   "PLC_a_HMI_Fila[6].Elemento[2].Estado" : Byte, 100 ms
   "PLC_a_HMI_Fila[6].Elemento[3].Figura" : Byte, 100 ms
   "PLC_a_HMI_Fila[6].Elemento[3].Offset_X" : Int, 100 ms
   "PLC_a_HMI_Fila[6].Elemento[3].Estado" : Byte, 100 ms
   "PLC_a_HMI_Fila[6].Elemento[4].Figura" : Byte, 100 ms
   "PLC_a_HMI_Fila[6].Elemento[4].Offset_X" : Int, 100 ms
   "PLC_a_HMI_Fila[6].Elemento[4].Estado" : Byte, 100 ms
   "PLC_a_HMI_Fila[6].Elemento[5].Figura" : Byte, 100 ms
   "PLC_a_HMI_Fila[6].Elemento[5].Offset_X" : Int, 100 ms
   "PLC_a_HMI_Fila[6].Elemento[5].Estado" : Byte, 100 ms
   "PLC_a_HMI_Fila[6].Elemento[6].Figura" : Byte, 100 ms
   "PLC_a_HMI_Fila[6].Elemento[6].Offset_X" : Int, 100 ms
   "PLC_a_HMI_Fila[6].Elemento[6].Estado" : Byte, 100 ms
   "PLC_a_HMI_Fila[6].Elemento[7].Figura" : Byte, 100 ms
   "PLC_a_HMI_Fila[6].Elemento[7].Offset_X" : Int, 100 ms
   "PLC_a_HMI_Fila[6].Elemento[7].Estado" : Byte, 100 ms
   "PLC_a_HMI_Fila[6].Elemento[8].Figura" : Byte, 100 ms
   "PLC_a_HMI_Fila[6].Elemento[8].Offset_X" : Int, 100 ms
   "PLC_a_HMI_Fila[6].Elemento[8].Estado" : Byte, 100 ms
   "PLC_a_HMI_Fila[6].Elemento[9].Figura" : Byte, 100 ms
   "PLC_a_HMI_Fila[6].Elemento[9].Offset_X" : Int, 100 ms
   "PLC_a_HMI_Fila[6].Elemento[9].Estado" : Byte, 100 ms
   "PLC_a_HMI_Fila[6].Elemento[10].Figura" : Byte, 100 ms
   "PLC_a_HMI_Fila[6].Elemento[10].Offset_X" : Int, 100 ms
   "PLC_a_HMI_Fila[6].Elemento[10].Estado" : Byte, 100 ms
   "PLC_a_HMI_Fila_Activa" : Byte, 1 s
   "DB_Animación_Figura_SEL" : Byte, 1 s
   "PLC_FechaHora" : Date_And_Time, 1 s
   "Proceso Empujador_Capa_Actual" : Byte, 1 s
   "DB_Receta_Actual_Nro_Capas_Pallet" : Byte, 1 s
   "Proceso Dosificador_Cant_Cajas" : Word, 1 s
   "DB_Receta_Actual_Nombre" : Array [0..49] of Char, 1 s
   "Proceso CargaPallet_Cant_Pallets" : DInt, 1 s
   "Proceso Empujador_Cant_Cajas" : DInt, 1 s
   "PLC a HMI_TRANSPORTES_Hab" : Bool, 1 s
   "PLC a HMI_Seg_Entrada_Envol" : Bool, 1 s
   "PLC a HMI_Seg_Salida_Envol" : Bool, 1 s
   "PLC a HMI_oTranspPall1" : Bool, 1 s
   "PLC a HMI_oTranspPall2" : Bool, 1 s
   "PLC a HMI_oTranspPall3" : Bool, 1 s
   "PLC a HMI_oTranspPall3Freno" : Bool, 1 s
   "PLC a HMI_oTranspPall4" : Bool, 1 s
   "PLC a HMI_oTranspPall5" : Bool, 1 s
   "PLC a HMI_iBrazoPos_Envolv" : Bool, 1 s
   "PLC a HMI_oHabilMovBrazo_Envol" : Bool, 1 s
   "PLC a HMI_iCartZonaSeg" : Bool, 1 s
   "PLC a HMI_iCartAplicado" : Bool, 1 s
   "PLC a HMI_iCartConAlarm" : Bool, 1 s
   "PLC a HMI_oTomarCartón" : Bool, 1 s
   "PLC a HMI_oAplicarCartón" : Bool, 1 s
   "PLC a HMI_oPaleZonaSeg" : Bool, 1 s
   "PLC a HMI_oPaleSinAlarm" : Bool, 1 s
   "FuncNormalAlterado" : Bool, 1 s
   "Confirmacion1" : Bool, internal
   "Confirmacion2" : Bool, internal

HMI tags "HMI_a_PLC"
   "HMI_Pls_Inc_Elem" : Bool, 1 s
   "HMI_Pls_Dec_Elem" : Bool, 1 s
   "HMI_Pls_Elem_Der" : Bool, 1 s
   "HMI_Pls_Elem_Izq" : Bool, 1 s
   "HMI_Pls_Inc_Fila" : Bool, 1 s
   "HMI_Pls_Dec_Fila" : Bool, 1 s
   "HMI_Pls_Fila_Sup" : Bool, 1 s
   "HMI_Pls_Fila_Inf" : Bool, 1 s
   "HMI_Pls_New_Fila" : Bool, 1 s
   "HMI_Pls_New_Elem" : Bool, 1 s
   "HMI_Pls_Kill_Elem" : Bool, 1 s
   "HMI_Pls_WR_Receta" : Bool, 1 s
   "HMI_Pls_RD_Receta" : Bool, 1 s
   "HMI_Imagen_Actual" : Word, 100 ms
   "HMI_Pls_Inc_Receta" : Bool, 1 s
   "HMI_Pls_Dec_Receta" : Bool, 1 s
   "HMI_Pls_Inc_Capa" : Bool, 1 s
   "HMI_Pls_Dec_Capa" : Bool, 1 s
   "HMI_Pls_Elem_+" : Bool, 1 s
   "HMI_Pls_Elem_-" : Bool, 1 s
   "HMI_Pls_CargarReceta" : Bool, 1 s
   "HMI_Pls_TerminarPallet" : Bool, 1 s
   "HMI_Pls_ResetPallets" : Bool, 1 s
   "HMI_Pls_ResetCajas" : Bool, 1 s
   "HMI_Pls_SalirImagenIni" : Bool, 1 s
   "HMI_Pls_MarMan_Ramp1" : Bool, 1 s
   "HMI_Pls_MarMan_Rol1" : Bool, 1 s
   "HMI_Pls_MarMan_Ramp2" : Bool, 1 s
   "HMI_Pls_MarMan_Rol2" : Bool, 1 s
   "HMI_Hab_Cartonero" : Bool, 1 s

discrete alarms
   1: '', class Grave, trigger "ALARMAS_1" bit 0
   2: '', class Grave, trigger "ALARMAS_1" bit 1
   3: '', class Grave, trigger "ALARMAS_1" bit 2
   4: '', class Grave, trigger "ALARMAS_1" bit 3
   5: '', class Grave, trigger "ALARMAS_1" bit 4
   6: '', class Grave, trigger "ALARMAS_1" bit 5
   7: '', class Grave, trigger "ALARMAS_1" bit 6
   8: '', class Grave, trigger "ALARMAS_1" bit 7
   9: '', class General, trigger "ALARMAS_1" bit 8
   10: '', class General, trigger "ALARMAS_1" bit 9
   11: '', class General, trigger "ALARMAS_1" bit 10
   12: '', class General, trigger "ALARMAS_1" bit 11
   13: '', class General, trigger "ALARMAS_1" bit 12
   14: '', class General, trigger "ALARMAS_1" bit 13
   15: '', class General, trigger "ALARMAS_1" bit 14
   16: '', class General, trigger "ALARMAS_1" bit 15
   17: '', class Transp. Cajas, trigger "ALARMAS_2" bit 0
   18: '', class Transp. Cajas, trigger "ALARMAS_2" bit 1
   19: '', class Transp. Cajas, trigger "ALARMAS_2" bit 2
   20: '', class Transp. Cajas, trigger "ALARMAS_2" bit 3
   21: '', class Transp. Cajas, trigger "ALARMAS_2" bit 4
   22: '', class Transp. Cajas, trigger "ALARMAS_2" bit 5
   23: '', class Transp. Cajas, trigger "ALARMAS_2" bit 6
   24: '', class Transp. Cajas, trigger "ALARMAS_2" bit 7
   25: '', class Transp. Cajas, trigger "ALARMAS_2" bit 8
   26: '', class Transp. Cajas, trigger "ALARMAS_2" bit 9
   27: '', class Transp. Cajas, trigger "ALARMAS_2" bit 10
   28: '', class Transp. Cajas, trigger "ALARMAS_2" bit 11
   29: '', class Transp. Cajas, trigger "ALARMAS_2" bit 12
   30: '', class Transp. Cajas, trigger "ALARMAS_2" bit 13
   31: '', class Transp. Cajas, trigger "ALARMAS_2" bit 14
   32: '', class Transp. Cajas, trigger "ALARMAS_2" bit 15
   33: '', class Dosificador, trigger "ALARMAS_3" bit 0
   34: '', class Dosificador, trigger "ALARMAS_3" bit 1
   35: '', class Dosificador, trigger "ALARMAS_3" bit 2
   36: '', class Dosificador, trigger "ALARMAS_3" bit 3
   37: '', class Dosificador, trigger "ALARMAS_3" bit 4
   38: '', class Dosificador, trigger "ALARMAS_3" bit 5
   39: '', class Dosificador, trigger "ALARMAS_3" bit 6
   40: '', class Dosificador, trigger "ALARMAS_3" bit 7
   41: '', class Dosificador, trigger "ALARMAS_3" bit 8
   42: '', class Dosificador, trigger "ALARMAS_3" bit 9
   43: '', class Dosificador, trigger "ALARMAS_3" bit 10
   44: '', class Dosificador, trigger "ALARMAS_3" bit 11
   45: '', class Dosificador, trigger "ALARMAS_3" bit 12
   46: '', class Dosificador, trigger "ALARMAS_3" bit 13
   47: '', class Dosificador, trigger "ALARMAS_3" bit 14
   48: '', class Dosificador, trigger "ALARMAS_3" bit 15
   49: '', class Carga Pallets, trigger "ALARMAS_4" bit 0
   50: '', class Carga Pallets, trigger "ALARMAS_4" bit 1
   51: '', class Carga Pallets, trigger "ALARMAS_4" bit 2
   52: '', class Carga Pallets, trigger "ALARMAS_4" bit 3
   53: '', class Carga Pallets, trigger "ALARMAS_4" bit 4
   54: '', class Carga Pallets, trigger "ALARMAS_4" bit 5
   55: '', class Carga Pallets, trigger "ALARMAS_4" bit 6
   56: '', class Carga Pallets, trigger "ALARMAS_4" bit 7
   57: '', class Carga Pallets, trigger "ALARMAS_4" bit 8
   58: '', class Carga Pallets, trigger "ALARMAS_4" bit 9
   59: '', class Carga Pallets, trigger "ALARMAS_4" bit 10
   60: '', class Carga Pallets, trigger "ALARMAS_4" bit 11
   61: '', class Carga Pallets, trigger "ALARMAS_4" bit 12
   62: '', class Carga Pallets, trigger "ALARMAS_4" bit 13
   63: '', class Carga Pallets, trigger "ALARMAS_4" bit 14
   64: '', class Carga Pallets, trigger "ALARMAS_4" bit 15
   65: '', class Carga Pallets, trigger "ALARMAS_5" bit 0
   66: '', class Carga Pallets, trigger "ALARMAS_5" bit 1
   67: '', class Carga Pallets, trigger "ALARMAS_5" bit 2
   68: '', class Carga Pallets, trigger "ALARMAS_5" bit 3
   69: '', class Carga Pallets, trigger "ALARMAS_5" bit 4
   70: '', class Carga Pallets, trigger "ALARMAS_5" bit 5
   71: '', class Carga Pallets, trigger "ALARMAS_5" bit 6
   72: '', class Carga Pallets, trigger "ALARMAS_5" bit 7
   73: '', class Carga Pallets, trigger "ALARMAS_5" bit 8
   74: '', class Carga Pallets, trigger "ALARMAS_5" bit 9
   75: '', class Carga Pallets, trigger "ALARMAS_5" bit 10
   76: '', class Carga Pallets, trigger "ALARMAS_5" bit 11
   77: '', class Carga Pallets, trigger "ALARMAS_5" bit 12
   78: '', class Carga Pallets, trigger "ALARMAS_5" bit 13
   79: '', class Carga Pallets, trigger "ALARMAS_5" bit 14
   80: '', class Carga Pallets, trigger "ALARMAS_5" bit 15
   81: '', class Transp. Pallets, trigger "ALARMAS_6" bit 0
   82: '', class Transp. Pallets, trigger "ALARMAS_6" bit 1
   83: '', class Transp. Pallets, trigger "ALARMAS_6" bit 2
   84: '', class Transp. Pallets, trigger "ALARMAS_6" bit 3
   85: '', class Transp. Pallets, trigger "ALARMAS_6" bit 4
   86: '', class Transp. Pallets, trigger "ALARMAS_6" bit 5
   87: '', class Transp. Pallets, trigger "ALARMAS_6" bit 6
   88: '', class Transp. Pallets, trigger "ALARMAS_6" bit 7
   89: '', class Transp. Pallets, trigger "ALARMAS_6" bit 8
   90: '', class Transp. Pallets, trigger "ALARMAS_6" bit 9
   91: '', class Transp. Pallets, trigger "ALARMAS_6" bit 10
   92: '', class Transp. Pallets, trigger "ALARMAS_6" bit 11
   93: '', class Transp. Pallets, trigger "ALARMAS_6" bit 12
   94: '', class Transp. Pallets, trigger "ALARMAS_6" bit 13
   95: '', class Transp. Pallets, trigger "ALARMAS_6" bit 14
   96: '', class Transp. Pallets, trigger "ALARMAS_6" bit 15
   97: '', class Mensaje, trigger "ALARMAS_7" bit 0
   98: '', class Mensaje, trigger "ALARMAS_7" bit 1
   99: '', class Mensaje, trigger "ALARMAS_7" bit 2
   100: '', class Mensaje, trigger "ALARMAS_7" bit 3
   101: '', class Mensaje, trigger "ALARMAS_7" bit 4
   102: '', class Mensaje, trigger "ALARMAS_7" bit 5
   103: '', class Mensaje, trigger "ALARMAS_7" bit 6
   104: '', class Mensaje, trigger "ALARMAS_7" bit 7
   105: '', class Mensaje, trigger "ALARMAS_7" bit 8
   106: '', class Mensaje, trigger "ALARMAS_7" bit 9
   107: '', class Mensaje, trigger "ALARMAS_7" bit 10
   108: '', class Mensaje, trigger "ALARMAS_7" bit 11
   109: '', class Mensaje, trigger "ALARMAS_7" bit 12
   110: '', class Mensaje, trigger "ALARMAS_7" bit 13
   111: '', class Mensaje, trigger "ALARMAS_7" bit 14
   112: '', class Mensaje, trigger "ALARMAS_7" bit 15
   113: '', class Dosificador, trigger "ALARMAS_8" bit 0
   114: '', class Dosificador, trigger "ALARMAS_8" bit 1
   115: '', class Dosificador, trigger "ALARMAS_8" bit 2
   116: '', class Dosificador, trigger "ALARMAS_8" bit 3
   117: '', class Dosificador, trigger "ALARMAS_8" bit 4
   118: '', class Dosificador, trigger "ALARMAS_8" bit 5
   119: '', class Dosificador, trigger "ALARMAS_8" bit 6
   120: '', class Dosificador, trigger "ALARMAS_8" bit 7
   121: '', class Dosificador, trigger "ALARMAS_8" bit 8
   122: '', class Dosificador, trigger "ALARMAS_8" bit 9
   123: '', class Dosificador, trigger "ALARMAS_8" bit 10
   124: '', class Dosificador, trigger "ALARMAS_8" bit 11
   125: '', class Dosificador, trigger "ALARMAS_8" bit 12
   126: '', class Dosificador, trigger "ALARMAS_8" bit 13
   127: '', class Dosificador, trigger "ALARMAS_8" bit 14
   128: '', class Dosificador bit 0

text list "Título": 0 ''; 1 ''; 2 ''; 3 ''; 20 ''; 11 ''; 32 ''; 33 ''; 70 ''; 71 ''; 72 ''; 73 ''; 21 ''; 30 ''; 22 ''; 14 ''; 34 ''; 40 ''; 41 ''; 42 ''; 31 ''

text list "Pistón": 0 ''; 1 ''

text list "Cant_cartones": 0 ''; 1 ''

screen "99_Elementos" 800x480
   Group "Group" at 725,14 size 62x50
   Group "Group_1" at 645,14 size 62x50
   Group "Group_2" at 565,14 size 62x50
   Group "Group_3" at 485,14 size 62x50
   Group "Group_4" at 405,14 size 62x50
   Group "Group_5" at 325,14 size 62x50
   Group "Group_6" at 245,14 size 62x50
   Group "Group_7" at 165,14 size 62x50
   Group "Group_8" at 85,14 size 62x50
   Group "Group_9" at 12,14 size 62x50
   Group "Group_10" at 12,70 size 62x50
   Group "Group_11" at 85,70 size 62x50
   Group "Group_12" at 165,70 size 62x50
   Group "Group_13" at 245,70 size 62x50
   Group "Group_14" at 325,70 size 62x50
   Group "Group_15" at 405,70 size 62x50
   Group "Group_16" at 485,70 size 62x50
   Group "Group_17" at 565,70 size 62x50
   Group "Group_18" at 645,70 size 62x50
   Group "Group_19" at 725,70 size 62x50
   Group "Group_20" at 725,126 size 62x50
   Group "Group_21" at 645,126 size 62x50
   Group "Group_22" at 565,126 size 62x50
   Group "Group_23" at 485,126 size 62x50
   Group "Group_24" at 405,126 size 62x50
   Group "Group_25" at 325,126 size 62x50
   Group "Group_26" at 245,126 size 62x50
   Group "Group_27" at 165,126 size 62x50
   Group "Group_28" at 85,126 size 62x50
   Group "Group_29" at 12,126 size 62x50
   Group "Group_30" at 12,182 size 62x50
   Group "Group_31" at 12,238 size 62x50
   Group "Group_32" at 12,294 size 62x50
   Group "Group_37" at 85,294 size 62x50
   Group "Group_38" at 85,238 size 62x50
   Group "Group_39" at 85,182 size 62x50
   Group "Group_40" at 165,182 size 62x50
   Group "Group_41" at 165,238 size 62x50
   Group "Group_42" at 165,294 size 62x50
   Group "Group_47" at 245,294 size 62x50
   Group "Group_48" at 245,238 size 62x50
   Group "Group_49" at 245,182 size 62x50
   Group "Group_50" at 325,182 size 62x50
   Group "Group_51" at 325,238 size 62x50
   Group "Group_52" at 325,294 size 62x50
   Group "Group_57" at 405,294 size 62x50
   Group "Group_58" at 405,238 size 62x50
   Group "Group_59" at 405,182 size 62x50
   Group "Group_60" at 485,182 size 62x50
   Group "Group_61" at 485,238 size 62x50
   Group "Group_62" at 485,294 size 62x50
   Group "Group_67" at 565,294 size 62x50
   Group "Group_68" at 565,238 size 62x50
   Group "Group_69" at 565,182 size 62x50
   Group "Group_70" at 645,182 size 62x50
   Group "Group_71" at 645,238 size 62x50
   Group "Group_72" at 645,294 size 62x50
   Group "Group_77" at 725,294 size 62x50
   Group "Group_78" at 725,238 size 62x50
   Group "Group_79" at 725,182 size 62x50

screen "98_Dibujo" 800x480
   Group "Group_33" at 362,384 size 122x84
   Group "Group" at 725,14 size 62x50
   Group "Group_19" at 725,38 size 62x50
   Group "Group_20" at 725,62 size 62x50
   Group "Group_79" at 725,86 size 62x50
   Group "Group_78" at 725,110 size 62x50
   Group "Group_77" at 725,134 size 62x50
   Group "Group_1" at 695,14 size 62x50
   Group "Group_18" at 695,38 size 62x50
   Group "Group_21" at 695,62 size 62x50
   Group "Group_70" at 695,86 size 62x50
   Group "Group_71" at 695,110 size 62x50
   Group "Group_72" at 695,134 size 62x50
   Group "Group_2" at 665,14 size 62x50
   Group "Group_17" at 665,38 size 62x50
   Group "Group_22" at 665,62 size 62x50
   Group "Group_69" at 665,86 size 62x50
   Group "Group_68" at 665,110 size 62x50
   Group "Group_67" at 665,134 size 62x50
   Group "Group_3" at 635,14 size 62x50
   Group "Group_16" at 635,38 size 62x50
   Group "Group_23" at 635,62 size 62x50
   Group "Group_60" at 635,86 size 62x50
   Group "Group_61" at 635,110 size 62x50
   Group "Group_62" at 635,134 size 62x50
   Group "Group_4" at 605,14 size 62x50
   Group "Group_15" at 605,38 size 62x50
   Group "Group_24" at 605,62 size 62x50
   Group "Group_59" at 605,86 size 62x50
   Group "Group_58" at 605,110 size 62x50
   Group "Group_57" at 605,134 size 62x50
   Group "Group_5" at 575,14 size 62x50
   Group "Group_14" at 575,38 size 62x50
   Group "Group_25" at 575,62 size 62x50
   Group "Group_50" at 575,86 size 62x50
   Group "Group_51" at 575,110 size 62x50
   Group "Group_52" at 575,134 size 62x50
   Group "Group_6" at 545,14 size 62x50
   Group "Group_13" at 545,38 size 62x50
   Group "Group_26" at 545,62 size 62x50
   Group "Group_49" at 545,86 size 62x50
   Group "Group_48" at 545,110 size 62x50
   Group "Group_47" at 545,134 size 62x50
   Group "Group_7" at 515,14 size 62x50
   Group "Group_12" at 515,38 size 62x50
   Group "Group_27" at 515,62 size 62x50
   Group "Group_40" at 515,86 size 62x50
   Group "Group_41" at 515,110 size 62x50
   Group "Group_42" at 515,134 size 62x50
   Group "Group_8" at 485,14 size 62x50
   Group "Group_11" at 485,38 size 62x50
   Group "Group_28" at 485,62 size 62x50
   Group "Group_39" at 485,86 size 62x50
   Group "Group_38" at 485,110 size 62x50
   Group "Group_37" at 485,134 size 62x50
   Group "Group_9" at 455,14 size 62x50
   Group "Group_10" at 455,38 size 62x50
   Group "Group_29" at 455,62 size 62x50
   Group "Group_30" at 455,86 size 62x50
   Group "Group_31" at 455,110 size 62x50
   Group "Group_32" at 455,134 size 62x50
   Button "Botón_4" at 80,288 size 80x64
   Button "Botón_6" at 160,352 size 80x64
   Button "Botón_7" at 0,352 size 80x64
   Button "Botón_9" at 80,416 size 80x64
   Button "Botón_1" at 362,384 size 122x84
   Button "Botón_2" at 0,288 size 80x64
   Button "Botón_3" at 160,416 size 80x64
   Button "Botón_5" at 80,352 size 80x64

screen "22_Recetas_Edit" 800x480, template "_Recetas_Editar"
   Group "Group" at 738,120 size 62x50
   Group "Group_19" at 738,144 size 62x50
   Group "Group_20" at 738,168 size 62x50
   Group "Group_79" at 738,192 size 62x50
   Group "Group_1" at 708,120 size 62x50
   Group "Group_18" at 708,144 size 62x50
   Group "Group_21" at 708,168 size 62x50
   Group "Group_70" at 708,192 size 62x50
   Group "Group_2" at 678,120 size 62x50
   Group "Group_17" at 678,144 size 62x50
   Group "Group_22" at 678,168 size 62x50
   Group "Group_69" at 678,192 size 62x50
   Group "Group_3" at 648,120 size 62x50
   Group "Group_16" at 648,144 size 62x50
   Group "Group_23" at 648,168 size 62x50
   Group "Group_60" at 648,192 size 62x50
   Group "Group_4" at 618,120 size 62x50
   Group "Group_15" at 618,144 size 62x50
   Group "Group_24" at 618,168 size 62x50
   Group "Group_59" at 618,192 size 62x50
   Group "Group_5" at 588,120 size 62x50
   Group "Group_14" at 588,144 size 62x50
   Group "Group_25" at 588,168 size 62x50
   Group "Group_50" at 588,192 size 62x50
   Group "Group_6" at 558,120 size 62x50
   Group "Group_13" at 558,144 size 62x50
   Group "Group_26" at 558,168 size 62x50
   Group "Group_49" at 558,192 size 62x50
   Group "Group_7" at 528,120 size 62x50
   Group "Group_12" at 528,144 size 62x50
   Group "Group_27" at 528,168 size 62x50
   Group "Group_40" at 528,192 size 62x50
   Group "Group_8" at 498,120 size 62x50
   Group "Group_11" at 498,144 size 62x50
   Group "Group_28" at 498,168 size 62x50
   Group "Group_39" at 498,192 size 62x50
   Group "Group_9" at 468,120 size 62x50
   Group "Group_10" at 468,144 size 62x50
   Group "Group_29" at 468,168 size 62x50
   Group "Group_30" at 468,192 size 62x50
   Button "Botón_12" at 22,224 size 160x80
   Button "Botón_13" at 22,314 size 160x80
   Group "Group_33" at 325,334 size 122x84
   Button "Botón_14" at 322,332 size 128x88
   Button "Botón_1" at 100,436 size 100x44
   Button "Botón_17" at 0,436 size 100x44
   Button "Botón_2" at 22,134 size 160x80
   TextField "Plantilla_Campo de texto_2" at 0,88 size 293x27
   IOField "Plantilla_Campo ES_2" at 368,88 size 432x30
   Button "Botón_3" at 548,336 size 122x84
   TextField "Campo de texto_1" at 298,228 size 338x78

screen "01_Online" 800x480, template "_Automático"
   Group "Group" at 540,92 size 62x50
   Group "Group_19" at 540,116 size 62x50
   Group "Group_20" at 540,140 size 62x50
   Group "Group_79" at 540,164 size 62x50
   Group "Group_1" at 510,92 size 62x50
   Group "Group_18" at 510,116 size 62x50
   Group "Group_21" at 510,140 size 62x50
   Group "Group_70" at 510,164 size 62x50
   Group "Group_2" at 480,92 size 62x50
   Group "Group_17" at 480,116 size 62x50
   Group "Group_22" at 480,140 size 62x50
   Group "Group_69" at 480,164 size 62x50
   Group "Group_3" at 450,92 size 62x50
   Group "Group_16" at 450,116 size 62x50
   Group "Group_23" at 450,140 size 62x50
   Group "Group_60" at 450,164 size 62x50
   Group "Group_4" at 420,92 size 62x50
   Group "Group_15" at 420,116 size 62x50
   Group "Group_24" at 420,140 size 62x50
   Group "Group_59" at 420,164 size 62x50
   Group "Group_5" at 390,92 size 62x50
   Group "Group_14" at 390,116 size 62x50
   Group "Group_25" at 390,140 size 62x50
   Group "Group_50" at 390,164 size 62x50
   Group "Group_6" at 360,92 size 62x50
   Group "Group_13" at 360,116 size 62x50
   Group "Group_26" at 360,140 size 62x50
   Group "Group_49" at 360,164 size 62x50
   Group "Group_7" at 330,92 size 62x50
   Group "Group_12" at 330,116 size 62x50
   Group "Group_27" at 330,140 size 62x50
   Group "Group_40" at 330,164 size 62x50
   Group "Group_8" at 300,92 size 62x50
   Group "Group_11" at 300,116 size 62x50
   Group "Group_28" at 300,140 size 62x50
   Group "Group_39" at 300,164 size 62x50
   Group "Group_9" at 270,92 size 62x50
   Group "Group_10" at 270,116 size 62x50
   Group "Group_29" at 270,140 size 62x50
   Group "Group_30" at 166,128 size 62x50
   Button "Botón_3" at 160,318 size 180x96
   Button "Botón_1" at 465,318 size 180x96
   TextField "Campo de texto_1" at 120,238 size 562x58
   Button "Botón_15" at 400,436 size 100x44
   Button "Botón_17" at 0,436 size 100x44
   TextField "Campo de texto_2" at 150,214 size 505x80

screen "20_Recetas" 800x480, template "_Recetas"
   TextField "Plantilla_Campo de texto_1" at 45,182 size 258x34
   TextField "Plantilla_Campo de texto_2" at 45,236 size 258x34
   TextField "Plantilla_Campo de texto_3" at 45,290 size 258x34
   IOField "Campo ES_1" at 318,182 size 432x34
   IOField "Campo ES_2" at 318,236 size 432x34
   IOField "Campo ES_3" at 318,290 size 432x34
   TextField "Plantilla_Campo de texto_4" at 45,130 size 258x34
   IOField "Campo ES_4" at 318,130 size 432x34
   TextField "Plantilla_Campo de texto_5" at 45,344 size 258x34
   Button "Botón_1" at 318,344 size 130x54
   Button "Botón_2" at 470,344 size 130x54
   Button "Botón_4" at 620,344 size 130x54

screen "02_Conteo" 800x480, template "_Automático"
   TextField "Plantilla_Campo de texto_2" at 65,214 size 391x25
   TextField "Plantilla_Campo de texto_3" at 65,310 size 392x25
   IOField "Campo ES_6" at 571,118 size 33x27
   IOField "Campo ES_7" at 657,118 size 33x27
   TextField "Plantilla_Campo de texto_6" at 65,118 size 396x25
   TextField "Plantilla_Campo de texto_7" at 621,118 size 25x25
   IOField "Campo ES_2" at 558,214 size 117x27
   IOField "Campo ES_3" at 558,310 size 117x27
   Button "Botón_1" at 489,152 size 136x48
   Button "Botón_2" at 639,152 size 136x48
   Button "Botón_3" at 535,248 size 200x48
   Button "Botón_4" at 535,344 size 200x48
   Button "Botón_13" at 100,436 size 100x44
   Button "Botón_5" at 60,376 size 96x32
   Button "Botón_6" at 155,376 size 96x32
   TextField "Campo de texto_1" at 219,130 size 343x118
   Button "Botón_7" at 264,223 size 96x32
   Button "Botón_8" at 424,223 size 96x32
   TextField "Campo de texto_2" at 219,130 size 343x118
   Button "Botón_9" at 264,223 size 96x32
   Button "Botón_10" at 424,223 size 96x32
   TextField "Campo de texto_3" at 62,349 size 186x23

screen "11_Alarmas" 800x480, template "_Alarmas"
   AlarmView "Plantilla_Visor de avisos_1" at 0,58 size 800x376

screen "32_Man_Empujador" 800x480, template "_Manual"
   TextField "Campo de texto_2" at 192,160 size 60x25
   TextField "Campo de texto_4" at 192,256 size 57x25
   TextField "Campo de texto_5" at 472,160 size 86x25
   TextField "Campo de texto_6" at 472,208 size 198x25
   TextField "Campo de texto_7" at 472,304 size 164x25
   TextField "Campo de texto_8" at 132,106 size 75x25
   TextField "Campo de texto_9" at 412,106 size 102x25
   TextField "Campo de texto_1" at 472,352 size 52x25
   TextField "Campo de texto_3" at 472,256 size 138x25
   Button "Botón_14" at 200,436 size 100x44

screen "33_Man_Plataforma" 800x480, template "_Manual"
   Switch "Interruptor_1" at 292,338 size 238x64
   TextField "Campo de texto_1" at 272,298 size 149x25
   TextField "Campo de texto_2" at 172,128 size 60x25
   TextField "Campo de texto_3" at 172,176 size 173x25
   TextField "Campo de texto_4" at 172,224 size 57x25
   TextField "Campo de texto_5" at 492,128 size 86x25
   TextField "Campo de texto_6" at 492,176 size 108x25
   TextField "Campo de texto_7" at 492,224 size 52x25
   TextField "Campo de texto_8" at 132,74 size 85x25
   TextField "Campo de texto_9" at 452,74 size 106x25
   Button "Botón_15" at 300,436 size 100x44

screen "14_eProC" 800x480
   Button "Botón_1" at 0,0 size 798x478
   GraphicView "Visor de gráficos_1" at 225,112 size 380x208

screen "70_Transp_Cajas" 800x480, template "_Transportes"
   Button "Botón_11" at 0,436 size 100x44
   TextField "Campo de texto_2" at 172,208 size 142x25
   TextField "Campo de texto_4" at 172,304 size 142x25
   TextField "Campo de texto_5" at 542,182 size 86x25
   TextField "Campo de texto_6" at 542,232 size 74x25
   TextField "Campo de texto_7" at 542,278 size 86x25
   TextField "Campo de texto_8" at 542,326 size 74x25
   TextField "Campo de texto_10" at 430,138 size 176x25
   TextField "Campo de texto_1" at 130,138 size 88x25

screen "73_Transp_Señales" 800x480, template "_Transportes"
   TextField "Campo de texto_1" at 92,142 size 121x25
   TextField "Campo de texto_2" at 92,180 size 147x25
   TextField "Campo de texto_3" at 92,220 size 140x25
   TextField "Campo de texto_5" at 472,142 size 152x25
   TextField "Campo de texto_6" at 472,180 size 84x25
   TextField "Campo de texto_7" at 472,220 size 124x25
   TextField "Campo de texto_4" at 50,102 size 221x25
   TextField "Campo de texto_8" at 430,102 size 226x25
   GraphicView "Visor de gráficos_1" at 18,178 size 28x30
   GraphicView "Visor de gráficos_2" at 18,140 size 28x30
   GraphicView "Visor de gráficos_3" at 18,218 size 28x30
   GraphicView "Visor de gráficos_4" at 398,140 size 28x30
   GraphicView "Visor de gráficos_5" at 398,178 size 28x30
   GraphicView "Visor de gráficos_6" at 398,218 size 28x30
   Button "Botón_15" at 400,436 size 100x44
   TextField "Campo de texto_9" at 92,302 size 216x25
   TextField "Campo de texto_10" at 92,340 size 222x25
   TextField "Campo de texto_11" at 92,380 size 154x25
   GraphicView "Visor de gráficos_8" at 18,300 size 28x30
   GraphicView "Visor de gráficos_9" at 18,378 size 28x30
   TextField "Campo de texto_12" at 472,302 size 133x25
   TextField "Campo de texto_13" at 472,340 size 138x25
   TextField "Campo de texto_14" at 472,380 size 220x25
   GraphicView "Visor de gráficos_10" at 398,300 size 28x30
   TextField "Campo de texto_15" at 472,264 size 239x25
   GraphicView "Visor de gráficos_13" at 398,262 size 28x30
   TextField "Campo de texto_16" at 50,260 size 125x25
   GraphicView "Visor de gráficos_7" at 18,340 size 28x30
   GraphicView "Visor de gráficos_11" at 398,340 size 28x30
   GraphicView "Visor de gráficos_12" at 398,380 size 28x30

screen "71_Transp_Pallets" 800x480, template "_Transportes"
   Button "Botón_7" at 100,436 size 100x44
   Group "Group_1" at 690,284 size 95x58
   Group "Group_2" at 588,284 size 95x58
   Group "Group_7" at 22,290 size 62x44
   TextField "Campo de texto_1" at 235,228 size 57x25
   TextField "Campo de texto_2" at 415,170 size 68x25
   TextField "Campo de texto_3" at 408,148 size 82x18
   TextField "Campo de texto_4" at 140,160 size 90x25
   TextField "Campo de texto_5" at 638,160 size 85x25
   Group "Group_6" at 135,290 size 62x44
   Group "Group_5" at 242,290 size 62x44
   Group "Group_4" at 440,290 size 62x44
   Group "Group_3" at 600,290 size 62x44
   Group "Group" at 705,290 size 62x44
   Group "Group_8" at 365,342 size 48x22
   TextField "Campo de texto_6" at 395,120 size 102x25

screen "21_Recetas" 800x480, template "_Recetas"
   Button "Botón_15" at 400,436 size 100x44
   Button "Botón_2" at 100,436 size 100x44
   Button "Botón_3" at 0,436 size 100x44
   Button "Botón_1" at 300,436 size 100x44
   TextField "Plantilla_Campo de texto_1" at 45,182 size 258x34
   TextField "Plantilla_Campo de texto_2" at 45,236 size 258x34
   TextField "Plantilla_Campo de texto_3" at 45,290 size 258x34
   IOField "Campo ES_1" at 318,182 size 432x34
   IOField "Campo ES_2" at 318,236 size 432x34
   IOField "Campo ES_3" at 318,290 size 432x34
   TextField "Plantilla_Campo de texto_4" at 45,130 size 258x34
   IOField "Campo ES_4" at 318,130 size 432x34

screen "30_Man_Palets" 800x480, template "_Manual"
   Button "Botón_11" at 100,436 size 100x44
   Button "Botón_2" at 622,352 size 138x48
   Button "Botón_3" at 495,64 size 138x48
   Button "Botón_1" at 292,64 size 138x48
   Button "Botón_4" at 165,352 size 138x48
   Button "Botón_5" at 25,352 size 138x48
   Group "Group_1" at 690,284 size 95x58
   Group "Group_2" at 588,284 size 95x58
   Group "Group_7" at 22,290 size 62x44
   TextField "Campo de texto_1" at 235,228 size 57x25
   TextField "Campo de texto_2" at 415,170 size 68x25
   TextField "Campo de texto_3" at 408,148 size 82x18
   TextField "Campo de texto_4" at 140,160 size 90x25
   TextField "Campo de texto_5" at 638,160 size 85x25
   Group "Group_6" at 135,290 size 62x44
   Group "Group_5" at 242,290 size 62x44
   Group "Group_4" at 440,290 size 62x44
   Group "Group_3" at 600,290 size 62x44
   Group "Group" at 705,290 size 62x44
   Group "Group_8" at 365,342 size 48x22
   TextField "Campo de texto_6" at 395,120 size 102x25

screen "34_Man_Ajustes" 800x480, template "_Manual"
   Button "Plantilla_Botón_1" at 280,128 size 240x64
   Button "Plantilla_Botón_2" at 280,210 size 240x64
   Button "Plantilla_Botón_3" at 280,288 size 240x64
   Button "Botón_16" at 600,436 size 100x44

screen "40_Ajus_Cinta" 800x480, template "_Ajustes"
   IOField "Campo ES_1" at 370,280 size 92x35
   IOField "Campo ES_2" at 370,232 size 92x35
   IOField "Campo ES_7" at 370,184 size 92x35
   TextField "Campo de texto_6" at 190,184 size 158x42
   TextField "Campo de texto_4" at 190,280 size 158x42

screen "41_Aju_Elevador" 800x480, template "_Ajustes"
   IOField "Campo ES_2" at 290,200 size 92x35
   TextField "Campo de texto_2" at 110,200 size 158x42
   IOField "Campo ES_3" at 290,248 size 92x35
   TextField "Campo de texto_3" at 110,248 size 158x42
   IOField "Campo ES_4" at 448,200 size 92x35
   IOField "Campo ES_5" at 448,248 size 92x35
   IOField "Campo ES_7" at 290,152 size 92x35
   IOField "Campo ES_1" at 290,296 size 92x35
   TextField "Campo de texto_1" at 315,100 size 64x31
   TextField "Campo de texto_6" at 110,152 size 158x42
   TextField "Campo de texto_4" at 110,296 size 158x42
   TextField "Campo de texto_5" at 475,100 size 65x31
   IOField "Campo ES_6" at 448,152 size 92x35
   IOField "Campo ES_8" at 448,296 size 92x35

screen "42_Aju_Empujador" 800x480, template "_Ajustes"
   IOField "Campo ES_2" at 290,200 size 92x35
   TextField "Campo de texto_2" at 110,200 size 158x42
   IOField "Campo ES_3" at 290,248 size 92x35
   TextField "Campo de texto_3" at 110,248 size 158x42
   IOField "Campo ES_4" at 448,200 size 92x35
   IOField "Campo ES_5" at 448,248 size 92x35
   IOField "Campo ES_6" at 448,296 size 92x35
   IOField "Campo ES_7" at 290,152 size 92x35
   IOField "Campo ES_1" at 290,296 size 92x35
   TextField "Campo de texto_1" at 285,100 size 107x31
   TextField "Campo de texto_6" at 110,152 size 158x42
   TextField "Campo de texto_4" at 110,296 size 158x42
   IOField "Campo ES_8" at 448,152 size 92x35
   TextField "Campo de texto_5" at 472,100 size 64x31

screen "31_Man_Cajas" 800x480, template "_Manual"
   Button "Botón_17" at 0,436 size 100x44
   Button "Botón_1" at 90,302 size 180x80
   Button "Botón_2" at 155,88 size 180x80
   Button "Botón_3" at 308,250 size 180x80
   Button "Botón_4" at 522,88 size 180x80
   TextField "Campo de texto_4" at 592,232 size 120x40
   TextField "Campo de texto_1" at 98,232 size 120x40

screen "23_Recetas_Param" 800x480, template "_Recetas"
   Button "Botón_1" at 100,436 size 100x44
   Button "Botón_17" at 0,436 size 100x44
   Button "Botón_2" at 400,436 size 100x44
   Button "Botón_3" at 300,436 size 100x44
   IOField "Campo ES_1" at 610,306 size 92x35
   IOField "Campo ES_2" at 610,258 size 92x35
   IOField "Campo ES_7" at 610,210 size 92x35
   TextField "Campo de texto_2" at 48,130 size 552x40
   IOField "Campo ES_4" at 608,130 size 132x40
   TextField "Campo de texto_3" at 48,258 size 552x40
   TextField "Campo de texto_1" at 48,210 size 552x40
   TextField "Campo de texto_5" at 48,306 size 552x40

Template "_Transportes" 800x480
   SymbolicIOField "Plantilla_Campo ES simbólico_1" at 0,0 size 800x58
   GraphicView "Plantilla_Visor de gráficos_1" at 2,2 size 135x56
   DateTimeField "Plantilla_Campo de fecha y hora_1" at 655,14 size 93x28
   TextField "Plantilla_Campo de texto_1" at 0,60 size 286x27
   Button "Botón_2" at 0,436 size 100x44
   Button "Botón_1" at 100,436 size 100x44
   Button "Botón_3" at 200,436 size 100x44
   Button "Botón_4" at 300,436 size 100x44
   Button "Botón_5" at 400,436 size 100x44
   Button "Botón_6" at 500,436 size 100x44
   Button "Botón_13" at 600,436 size 100x44
   Button "Botón_14" at 700,436 size 100x44
   IOField "Campo ES_1" at 286,60 size 514x27

Template "_Manual" 800x480
   SymbolicIOField "Plantilla_Campo ES simbólico_1" at 0,0 size 800x58
   GraphicView "Plantilla_Visor de gráficos_1" at 2,2 size 135x56
   DateTimeField "Plantilla_Campo de fecha y hora_1" at 655,14 size 93x28
   Button "Botón_2" at 0,436 size 100x44
   Button "Botón_1" at 100,436 size 100x44
   Button "Botón_3" at 200,436 size 100x44
   Button "Botón_4" at 300,436 size 100x44
   Button "Botón_5" at 400,436 size 100x44
   Button "Botón_6" at 500,436 size 100x44
   Button "Botón_7" at 600,436 size 100x44
   Button "Botón_8" at 700,436 size 100x44

Template "_Alarmas" 800x480
   SymbolicIOField "Plantilla_Campo ES simbólico_1" at 0,0 size 800x58
   GraphicView "Plantilla_Visor de gráficos_1" at 2,2 size 135x56
   DateTimeField "Plantilla_Campo de fecha y hora_1" at 655,14 size 93x28
   Button "Botón_2" at 0,436 size 100x44
   Button "Botón_1" at 100,436 size 100x44
   Button "Botón_3" at 200,436 size 100x44
   Button "Botón_4" at 300,436 size 100x44
   Button "Botón_5" at 400,436 size 100x44
   Button "Botón_6" at 500,436 size 100x44
   Button "Botón_13" at 600,436 size 100x44
   Button "Botón_14" at 700,436 size 100x44
   Button "Botón_7" at 500,436 size 100x44

Template "_Automático" 800x480
   SymbolicIOField "Plantilla_Campo ES simbólico_1" at 0,0 size 800x58
   GraphicView "Plantilla_Visor de gráficos_1" at 2,2 size 135x56
   DateTimeField "Plantilla_Campo de fecha y hora_1" at 655,14 size 93x28
   TextField "Plantilla_Campo de texto_1" at 0,60 size 286x27
   IOField "Campo ES_1" at 286,60 size 514x27
   Button "Botón_2" at 0,436 size 100x44
   Button "Botón_1" at 100,436 size 100x44
   Button "Botón_3" at 200,436 size 100x44
   Button "Botón_4" at 300,436 size 100x44
   Button "Botón_5" at 400,436 size 100x44
   Button "Botón_6" at 500,436 size 100x44
   Button "Botón_7" at 600,436 size 100x44
   Button "Botón_8" at 700,436 size 100x44

Template "_Recetas" 800x480
   SymbolicIOField "Plantilla_Campo ES simbólico_1" at 0,0 size 800x58
   GraphicView "Plantilla_Visor de gráficos_1" at 2,2 size 135x56
   DateTimeField "Plantilla_Campo de fecha y hora_1" at 655,14 size 93x28
   TextField "Plantilla_Campo de texto_1" at 0,60 size 286x27
   Button "Botón_2" at 0,436 size 100x44
   Button "Botón_1" at 100,436 size 100x44
   Button "Botón_3" at 200,436 size 100x44
   Button "Botón_4" at 300,436 size 100x44
   Button "Botón_5" at 400,436 size 100x44
   Button "Botón_6" at 500,436 size 100x44
   Button "Botón_7" at 600,436 size 100x44
   Button "Botón_8" at 700,436 size 100x44
   IOField "Campo ES_1" at 286,60 size 514x27

Template "_Recetas_Editar" 800x480
   SymbolicIOField "Plantilla_Campo ES simbólico_1" at 0,0 size 800x58
   GraphicView "Plantilla_Visor de gráficos_1" at 2,2 size 135x56
   DateTimeField "Plantilla_Campo de fecha y hora_1" at 655,14 size 93x28
   TextField "Plantilla_Campo de texto_1" at 0,58 size 281x27
   IOField "Plantilla_Campo ES_1" at 360,58 size 440x30
   Button "Botón_2" at 0,436 size 100x44
   Button "Botón_1" at 100,436 size 100x44
   Button "Botón_3" at 200,436 size 100x44
   Button "Botón_4" at 300,436 size 100x44
   Button "Botón_5" at 400,436 size 100x44
   Button "Botón_6" at 500,436 size 100x44
   Button "Botón_7" at 600,436 size 100x44
   Button "Botón_8" at 700,436 size 100x44

Template "_Ajustes" 800x480
   SymbolicIOField "Plantilla_Campo ES simbólico_1" at 0,0 size 800x58
   GraphicView "Plantilla_Visor de gráficos_1" at 2,2 size 135x56
   DateTimeField "Plantilla_Campo de fecha y hora_1" at 655,14 size 93x28
   Button "Botón_2" at 0,436 size 100x44
   Button "Botón_1" at 100,436 size 100x44
   Button "Botón_3" at 200,436 size 100x44
   Button "Botón_4" at 300,436 size 100x44
   Button "Botón_5" at 400,436 size 100x44
   Button "Botón_6" at 500,436 size 100x44
   Button "Botón_7" at 600,436 size 100x44
   Button "Botón_8" at 700,436 size 100x44

screen "20_Recetas_NO SE USA TEMPOR" 800x480, template "_Recetas"
   TextField "Plantilla_Campo de texto_1" at 45,182 size 258x34
   TextField "Plantilla_Campo de texto_2" at 45,236 size 258x34
   TextField "Plantilla_Campo de texto_3" at 45,290 size 258x34
   IOField "Campo ES_1" at 318,182 size 432x34
   IOField "Campo ES_2" at 318,236 size 432x34
   IOField "Campo ES_3" at 318,290 size 432x34
   TextField "Plantilla_Campo de texto_4" at 45,130 size 258x34
   IOField "Campo ES_4" at 318,130 size 432x34
   TextField "Plantilla_Campo de texto_5" at 45,344 size 258x34
   Button "Botón_1" at 318,344 size 130x54
   Button "Botón_2" at 470,344 size 130x54
   Button "Botón_4" at 620,344 size 130x54

screen "35_HabilitacionFallas" 800x480, template "_Alarmas"
   TextField "Campo de texto_1" at 52,107 size 79x27
   TextField "Campo de texto_2" at 76,146 size 128x27
   TextField "Campo de texto_3" at 83,202 size 121x27
   TextField "Campo de texto_4" at 83,258 size 121x27
   Switch "Interruptor_1" at 216,135 size 88x45
   Switch "Interruptor_2" at 216,191 size 88x45
   Switch "Interruptor_3" at 216,247 size 88x45
   IOField "Campo ES_1" at 510,236 size 180x56
   TextField "Campo de texto_5" at 500,115 size 207x27
   TextField "Campo de texto_6" at 480,155 size 250x27
   TextField "Campo de texto_7" at 480,187 size 240x27
*)